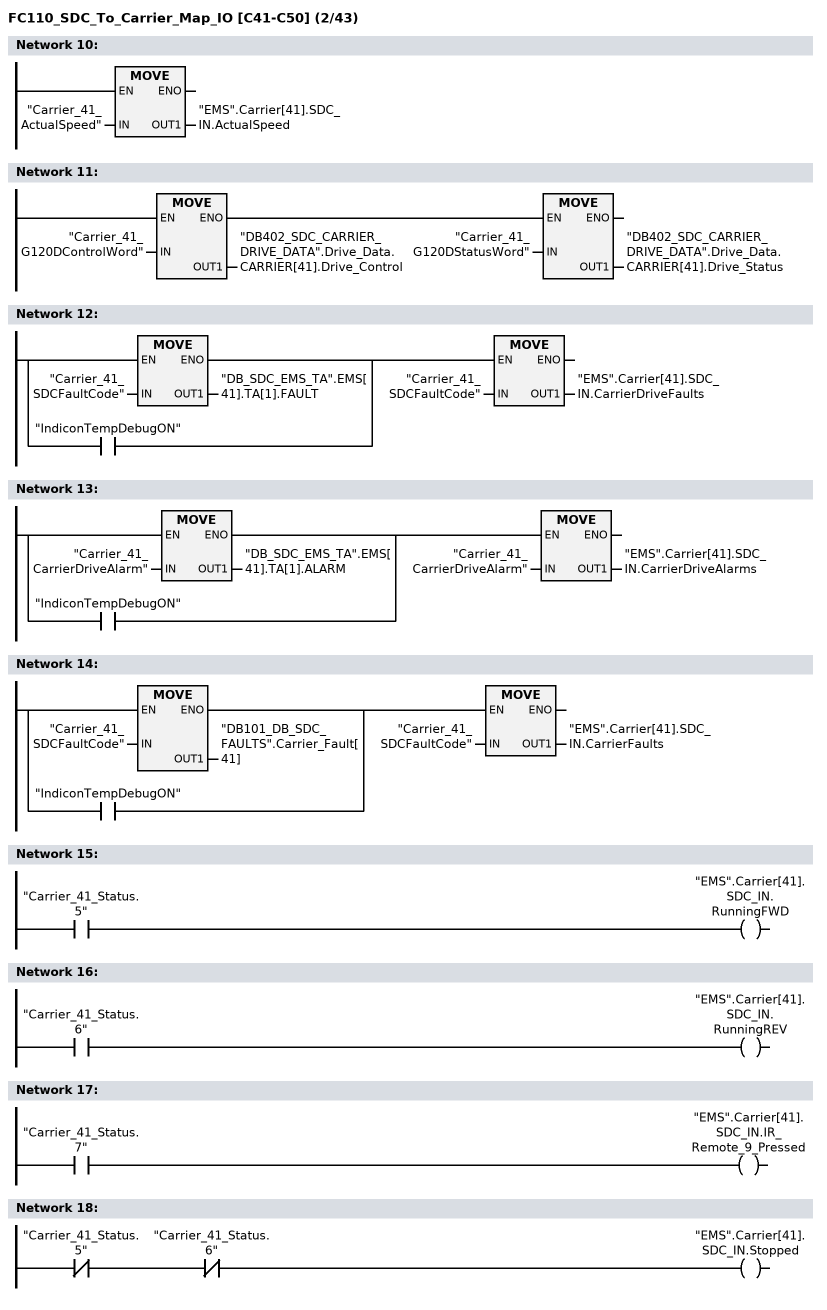
   RUNG wire#powerrail
      Move(in := "Carrier_41_ActualSpeed", out1 => "EMS".Carrier[41].SDC_IN.ActualSpeed)
   END_RUNG
   // the same network as SCL:
   "EMS".Carrier[41].SDC_IN.ActualSpeed := "Carrier_41_ActualSpeed";
END_REGION

REGION Network 11
   RUNG wire#powerrail
      Move(in := "Carrier_41_G120DControlWord", out1 => "DB402_SDC_CARRIER_DRIVE_DATA".Drive_Data.CARRIER[41].Drive_Control)
      Move(in := "Carrier_41_G120DStatusWord", out1 => "DB402_SDC_CARRIER_DRIVE_DATA".Drive_Data.CARRIER[41].Drive_Status)
   END_RUNG
   // the same network as SCL:
   "DB402_SDC_CARRIER_DRIVE_DATA".Drive_Data.CARRIER[41].Drive_Control := "Carrier_41_G120DControlWord";
   "DB402_SDC_CARRIER_DRIVE_DATA".Drive_Data.CARRIER[41].Drive_Status := "Carrier_41_G120DStatusWord";
END_REGION

REGION Network 12
   RUNG wire#powerrail
      Move(in := "Carrier_41_SDCFaultCode", out1 => "DB_SDC_EMS_TA".EMS[41].TA[1].FAULT)
      wire#w1
      Move(in := "Carrier_41_SDCFaultCode", out1 => "EMS".Carrier[41].SDC_IN.CarrierDriveFaults)
   END_RUNG
   RUNG wire#powerrail
      Contact( "IndiconTempDebugON" )
   END_RUNG wire#w1
   // the same network as SCL:
   "DB_SDC_EMS_TA".EMS[41].TA[1].FAULT := "Carrier_41_SDCFaultCode";
   IF TRUE OR "IndiconTempDebugON" THEN
       "EMS".Carrier[41].SDC_IN.CarrierDriveFaults := "Carrier_41_SDCFaultCode";
   END_IF;
END_REGION

REGION Network 13
   RUNG wire#powerrail
      Move(in := "Carrier_41_CarrierDriveAlarm", out1 => "DB_SDC_EMS_TA".EMS[41].TA[1].ALARM)
      wire#w1
      Move(in := "Carrier_41_CarrierDriveAlarm", out1 => "EMS".Carrier[41].SDC_IN.CarrierDriveAlarms)
   END_RUNG
   RUNG wire#powerrail
      Contact( "IndiconTempDebugON" )
   END_RUNG wire#w1
   // the same network as SCL:
   "DB_SDC_EMS_TA".EMS[41].TA[1].ALARM := "Carrier_41_CarrierDriveAlarm";
   IF TRUE OR "IndiconTempDebugON" THEN
       "EMS".Carrier[41].SDC_IN.CarrierDriveAlarms := "Carrier_41_CarrierDriveAlarm";
   END_IF;
END_REGION

REGION Network 14
   RUNG wire#powerrail
      Move(in := "Carrier_41_SDCFaultCode", out1 => "DB101_DB_SDC_FAULTS".Carrier_Fault[41])
      wire#w1
      Move(in := "Carrier_41_SDCFaultCode", out1 => "EMS".Carrier[41].SDC_IN.CarrierFaults)
   END_RUNG
   RUNG wire#powerrail
      Contact( "IndiconTempDebugON" )
   END_RUNG wire#w1
   // the same network as SCL:
   "DB101_DB_SDC_FAULTS".Carrier_Fault[41] := "Carrier_41_SDCFaultCode";
   IF TRUE OR "IndiconTempDebugON" THEN
       "EMS".Carrier[41].SDC_IN.CarrierFaults := "Carrier_41_SDCFaultCode";
   END_IF;
END_REGION

REGION Network 15
   RUNG wire#powerrail
      Contact( "Carrier_41_Status.5" )
      Coil( "EMS".Carrier[41].SDC_IN.RunningFWD )
   END_RUNG
   // the same network as SCL:
   "EMS".Carrier[41].SDC_IN.RunningFWD := "Carrier_41_Status.5";
END_REGION

REGION Network 16
   RUNG wire#powerrail
      Contact( "Carrier_41_Status.6" )
      Coil( "EMS".Carrier[41].SDC_IN.RunningREV )
   END_RUNG
   // the same network as SCL:
   "EMS".Carrier[41].SDC_IN.RunningREV := "Carrier_41_Status.6";
END_REGION

REGION Network 17
   RUNG wire#powerrail
      Contact( "Carrier_41_Status.7" )
      Coil( "EMS".Carrier[41].SDC_IN.IR_Remote_9_Pressed )
   END_RUNG
   // the same network as SCL:
   "EMS".Carrier[41].SDC_IN.IR_Remote_9_Pressed := "Carrier_41_Status.7";
END_REGION

REGION Network 18
   RUNG wire#powerrail
      I_Contact( "Carrier_41_Status.5" )
      I_Contact( "Carrier_41_Status.6" )
      Coil( "EMS".Carrier[41].SDC_IN.Stopped )
   END_RUNG
   // the same network as SCL:
   "EMS".Carrier[41].SDC_IN.Stopped := NOT "Carrier_41_Status.5" AND NOT "Carrier_41_Status.6";
END_REGION

REGION Network 19
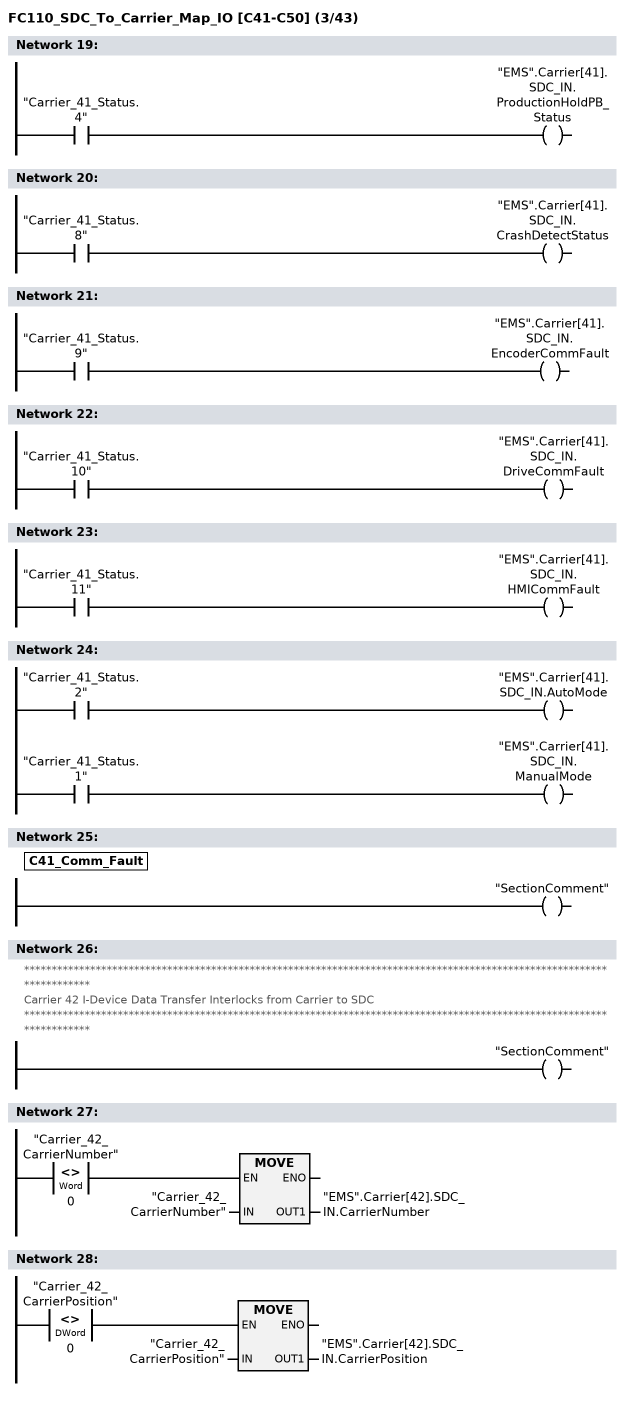
   RUNG wire#powerrail
      Contact( "Carrier_41_Status.4" )
      Coil( "EMS".Carrier[41].SDC_IN.ProductionHoldPB_Status )
   END_RUNG
   // the same network as SCL:
   "EMS".Carrier[41].SDC_IN.ProductionHoldPB_Status := "Carrier_41_Status.4";
END_REGION

REGION Network 20
   RUNG wire#powerrail
      Contact( "Carrier_41_Status.8" )
      Coil( "EMS".Carrier[41].SDC_IN.CrashDetectStatus )
   END_RUNG
   // the same network as SCL:
   "EMS".Carrier[41].SDC_IN.CrashDetectStatus := "Carrier_41_Status.8";
END_REGION

REGION Network 21
   RUNG wire#powerrail
      Contact( "Carrier_41_Status.9" )
      Coil( "EMS".Carrier[41].SDC_IN.EncoderCommFault )
   END_RUNG
   // the same network as SCL:
   "EMS".Carrier[41].SDC_IN.EncoderCommFault := "Carrier_41_Status.9";
END_REGION

REGION Network 22
   RUNG wire#powerrail
      Contact( "Carrier_41_Status.10" )
      Coil( "EMS".Carrier[41].SDC_IN.DriveCommFault )
   END_RUNG
   // the same network as SCL:
   "EMS".Carrier[41].SDC_IN.DriveCommFault := "Carrier_41_Status.10";
END_REGION

REGION Network 23
   RUNG wire#powerrail
      Contact( "Carrier_41_Status.11" )
      Coil( "EMS".Carrier[41].SDC_IN.HMICommFault )
   END_RUNG
   // the same network as SCL:
   "EMS".Carrier[41].SDC_IN.HMICommFault := "Carrier_41_Status.11";
END_REGION

REGION Network 24
   RUNG wire#powerrail
      Contact( "Carrier_41_Status.2" )
      Coil( "EMS".Carrier[41].SDC_IN.AutoMode )
   END_RUNG
   RUNG wire#powerrail
      Contact( "Carrier_41_Status.1" )
      Coil( "EMS".Carrier[41].SDC_IN.ManualMode )
   END_RUNG
   // the same network as SCL:
   "EMS".Carrier[41].SDC_IN.AutoMode := "Carrier_41_Status.2";
   "EMS".Carrier[41].SDC_IN.ManualMode := "Carrier_41_Status.1";
END_REGION

REGION Network 25
   Label( C41_Comm_Fault )
   RUNG wire#powerrail
      Coil( "SectionComment" )
   END_RUNG
   // the same network as SCL:
   C41_Comm_Fault:
   "SectionComment" := TRUE;
END_REGION

REGION Network 26
   // **********************************************************************************************************************
   // 
   // Carrier 42 I-Device Data Transfer Interlocks from Carrier to SDC
   // 
   // **********************************************************************************************************************
   RUNG wire#powerrail
      Coil( "SectionComment" )
   END_RUNG
   // the same network as SCL:
   "SectionComment" := TRUE;
END_REGION

REGION Network 27
   RUNG wire#powerrail
      { S7_Templates := "SrcType := Word" } NE_Contact(in1 := "Carrier_42_CarrierNumber", in2 := 0)
      Move(in := "Carrier_42_CarrierNumber", out1 => "EMS".Carrier[42].SDC_IN.CarrierNumber)
   END_RUNG
   // the same network as SCL:
   IF "Carrier_42_CarrierNumber" <> 0 THEN
       "EMS".Carrier[42].SDC_IN.CarrierNumber := "Carrier_42_CarrierNumber";
   END_IF;
END_REGION

REGION Network 28
   RUNG wire#powerrail
      { S7_Templates := "SrcType := DWord" } NE_Contact(in1 := "Carrier_42_CarrierPosition", in2 := 0)
      Move(in := "Carrier_42_CarrierPosition", out1 => "EMS".Carrier[42].SDC_IN.CarrierPosition)
   END_RUNG
   // the same network as SCL:
   IF "Carrier_42_CarrierPosition" <> 0 THEN
       "EMS".Carrier[42].SDC_IN.CarrierPosition := "Carrier_42_CarrierPosition";
   END_IF;
END_REGION

REGION Network 29
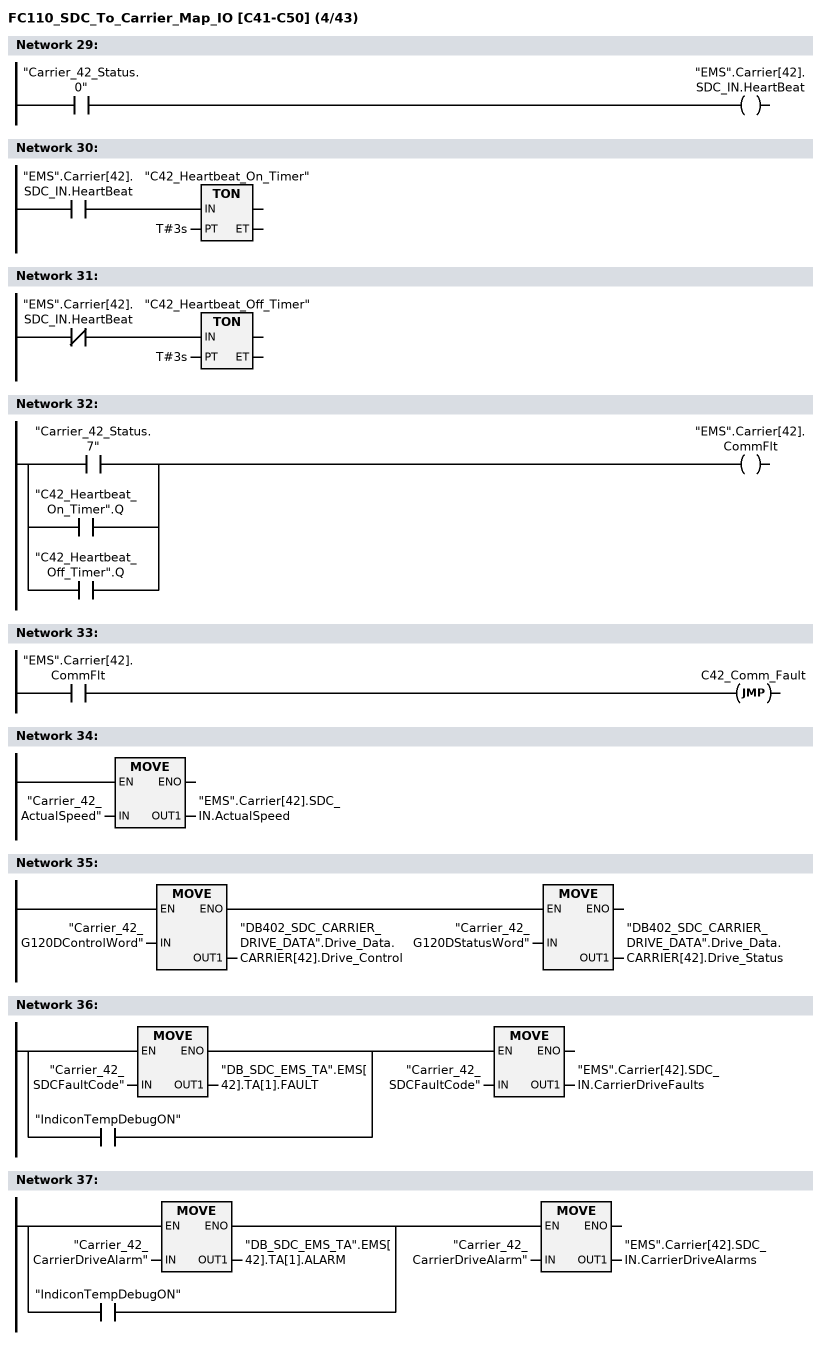
   RUNG wire#powerrail
      Contact( "Carrier_42_Status.0" )
      Coil( "EMS".Carrier[42].SDC_IN.HeartBeat )
   END_RUNG
   // the same network as SCL:
   "EMS".Carrier[42].SDC_IN.HeartBeat := "Carrier_42_Status.0";
END_REGION

REGION Network 30
   "C42_Heartbeat_On_Timer".TON(IN := "EMS".Carrier[42].SDC_IN.HeartBeat, PT := T#3s);
END_REGION

REGION Network 31
   "C42_Heartbeat_Off_Timer".TON(IN := NOT "EMS".Carrier[42].SDC_IN.HeartBeat, PT := T#3s);
END_REGION

REGION Network 32
   RUNG wire#powerrail
      Contact( "Carrier_42_Status.7" )
      wire#w1
      Coil( "EMS".Carrier[42].CommFlt )
   END_RUNG
   RUNG wire#powerrail
      Contact( "C42_Heartbeat_On_Timer".Q )
   END_RUNG wire#w1
   RUNG wire#powerrail
      Contact( "C42_Heartbeat_Off_Timer".Q )
   END_RUNG wire#w1
   // the same network as SCL:
   "EMS".Carrier[42].CommFlt := "Carrier_42_Status.7" OR "C42_Heartbeat_On_Timer".Q OR "C42_Heartbeat_Off_Timer".Q;
END_REGION

REGION Network 33
   RUNG wire#powerrail
      Contact( "EMS".Carrier[42].CommFlt )
      JumpCoil( C42_Comm_Fault )
   END_RUNG
   // the same network as SCL:
   IF "EMS".Carrier[42].CommFlt THEN GOTO C42_Comm_Fault; END_IF;
END_REGION

REGION Network 34
   RUNG wire#powerrail
      Move(in := "Carrier_42_ActualSpeed", out1 => "EMS".Carrier[42].SDC_IN.ActualSpeed)
   END_RUNG
   // the same network as SCL:
   "EMS".Carrier[42].SDC_IN.ActualSpeed := "Carrier_42_ActualSpeed";
END_REGION

REGION Network 35
   RUNG wire#powerrail
      Move(in := "Carrier_42_G120DControlWord", out1 => "DB402_SDC_CARRIER_DRIVE_DATA".Drive_Data.CARRIER[42].Drive_Control)
      Move(in := "Carrier_42_G120DStatusWord", out1 => "DB402_SDC_CARRIER_DRIVE_DATA".Drive_Data.CARRIER[42].Drive_Status)
   END_RUNG
   // the same network as SCL:
   "DB402_SDC_CARRIER_DRIVE_DATA".Drive_Data.CARRIER[42].Drive_Control := "Carrier_42_G120DControlWord";
   "DB402_SDC_CARRIER_DRIVE_DATA".Drive_Data.CARRIER[42].Drive_Status := "Carrier_42_G120DStatusWord";
END_REGION

REGION Network 36
   RUNG wire#powerrail
      Move(in := "Carrier_42_SDCFaultCode", out1 => "DB_SDC_EMS_TA".EMS[42].TA[1].FAULT)
      wire#w1
      Move(in := "Carrier_42_SDCFaultCode", out1 => "EMS".Carrier[42].SDC_IN.CarrierDriveFaults)
   END_RUNG
   RUNG wire#powerrail
      Contact( "IndiconTempDebugON" )
   END_RUNG wire#w1
   // the same network as SCL:
   "DB_SDC_EMS_TA".EMS[42].TA[1].FAULT := "Carrier_42_SDCFaultCode";
   IF TRUE OR "IndiconTempDebugON" THEN
       "EMS".Carrier[42].SDC_IN.CarrierDriveFaults := "Carrier_42_SDCFaultCode";
   END_IF;
END_REGION

REGION Network 37
   RUNG wire#powerrail
      Move(in := "Carrier_42_CarrierDriveAlarm", out1 => "DB_SDC_EMS_TA".EMS[42].TA[1].ALARM)
      wire#w1
      Move(in := "Carrier_42_CarrierDriveAlarm", out1 => "EMS".Carrier[42].SDC_IN.CarrierDriveAlarms)
   END_RUNG
   RUNG wire#powerrail
      Contact( "IndiconTempDebugON" )
   END_RUNG wire#w1
   // the same network as SCL:
   "DB_SDC_EMS_TA".EMS[42].TA[1].ALARM := "Carrier_42_CarrierDriveAlarm";
   IF TRUE OR "IndiconTempDebugON" THEN
       "EMS".Carrier[42].SDC_IN.CarrierDriveAlarms := "Carrier_42_CarrierDriveAlarm";
   END_IF;
END_REGION

REGION Network 38
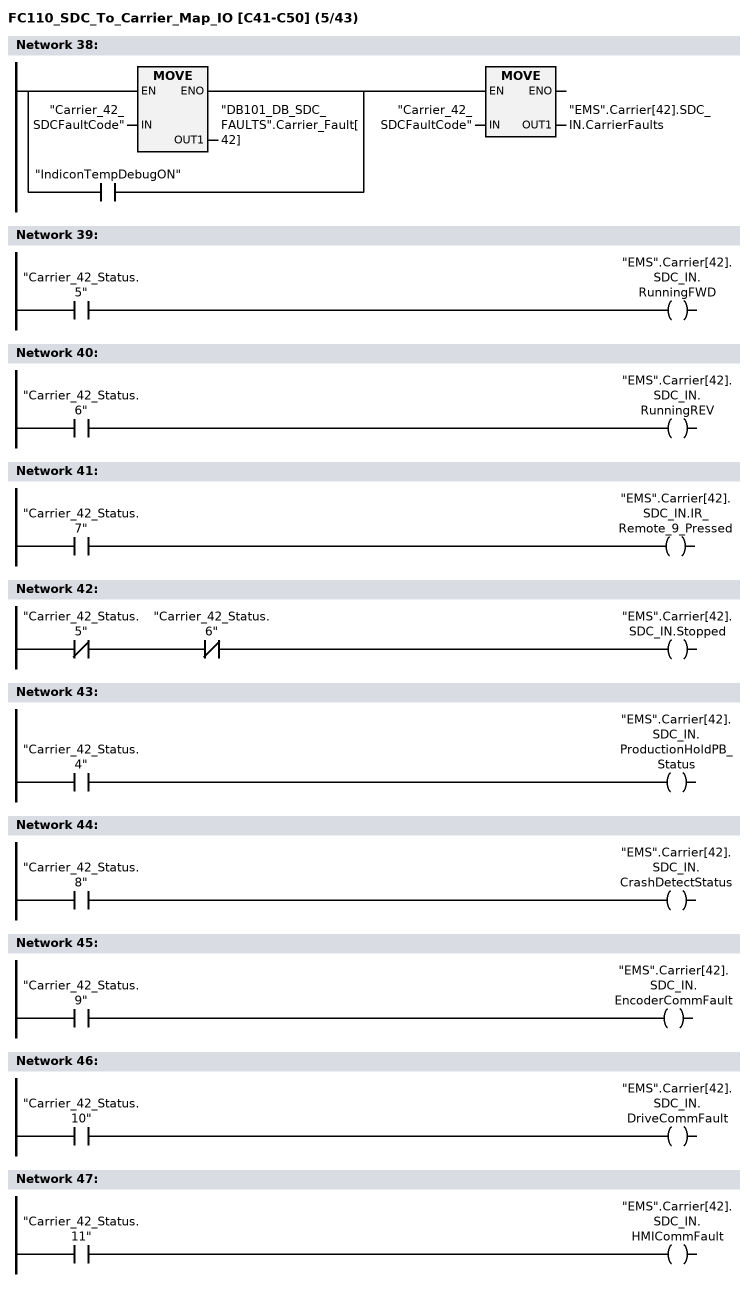
   RUNG wire#powerrail
      Move(in := "Carrier_42_SDCFaultCode", out1 => "DB101_DB_SDC_FAULTS".Carrier_Fault[42])
      wire#w1
      Move(in := "Carrier_42_SDCFaultCode", out1 => "EMS".Carrier[42].SDC_IN.CarrierFaults)
   END_RUNG
   RUNG wire#powerrail
      Contact( "IndiconTempDebugON" )
   END_RUNG wire#w1
   // the same network as SCL:
   "DB101_DB_SDC_FAULTS".Carrier_Fault[42] := "Carrier_42_SDCFaultCode";
   IF TRUE OR "IndiconTempDebugON" THEN
       "EMS".Carrier[42].SDC_IN.CarrierFaults := "Carrier_42_SDCFaultCode";
   END_IF;
END_REGION

REGION Network 39
   RUNG wire#powerrail
      Contact( "Carrier_42_Status.5" )
      Coil( "EMS".Carrier[42].SDC_IN.RunningFWD )
   END_RUNG
   // the same network as SCL:
   "EMS".Carrier[42].SDC_IN.RunningFWD := "Carrier_42_Status.5";
END_REGION

REGION Network 40
   RUNG wire#powerrail
      Contact( "Carrier_42_Status.6" )
      Coil( "EMS".Carrier[42].SDC_IN.RunningREV )
   END_RUNG
   // the same network as SCL:
   "EMS".Carrier[42].SDC_IN.RunningREV := "Carrier_42_Status.6";
END_REGION

REGION Network 41
   RUNG wire#powerrail
      Contact( "Carrier_42_Status.7" )
      Coil( "EMS".Carrier[42].SDC_IN.IR_Remote_9_Pressed )
   END_RUNG
   // the same network as SCL:
   "EMS".Carrier[42].SDC_IN.IR_Remote_9_Pressed := "Carrier_42_Status.7";
END_REGION

REGION Network 42
   RUNG wire#powerrail
      I_Contact( "Carrier_42_Status.5" )
      I_Contact( "Carrier_42_Status.6" )
      Coil( "EMS".Carrier[42].SDC_IN.Stopped )
   END_RUNG
   // the same network as SCL:
   "EMS".Carrier[42].SDC_IN.Stopped := NOT "Carrier_42_Status.5" AND NOT "Carrier_42_Status.6";
END_REGION

REGION Network 43
   RUNG wire#powerrail
      Contact( "Carrier_42_Status.4" )
      Coil( "EMS".Carrier[42].SDC_IN.ProductionHoldPB_Status )
   END_RUNG
   // the same network as SCL:
   "EMS".Carrier[42].SDC_IN.ProductionHoldPB_Status := "Carrier_42_Status.4";
END_REGION

REGION Network 44
   RUNG wire#powerrail
      Contact( "Carrier_42_Status.8" )
      Coil( "EMS".Carrier[42].SDC_IN.CrashDetectStatus )
   END_RUNG
   // the same network as SCL:
   "EMS".Carrier[42].SDC_IN.CrashDetectStatus := "Carrier_42_Status.8";
END_REGION

REGION Network 45
   RUNG wire#powerrail
      Contact( "Carrier_42_Status.9" )
      Coil( "EMS".Carrier[42].SDC_IN.EncoderCommFault )
   END_RUNG
   // the same network as SCL:
   "EMS".Carrier[42].SDC_IN.EncoderCommFault := "Carrier_42_Status.9";
END_REGION

REGION Network 46
   RUNG wire#powerrail
      Contact( "Carrier_42_Status.10" )
      Coil( "EMS".Carrier[42].SDC_IN.DriveCommFault )
   END_RUNG
   // the same network as SCL:
   "EMS".Carrier[42].SDC_IN.DriveCommFault := "Carrier_42_Status.10";
END_REGION

REGION Network 47
   RUNG wire#powerrail
      Contact( "Carrier_42_Status.11" )
      Coil( "EMS".Carrier[42].SDC_IN.HMICommFault )
   END_RUNG
   // the same network as SCL:
   "EMS".Carrier[42].SDC_IN.HMICommFault := "Carrier_42_Status.11";
END_REGION

REGION Network 48
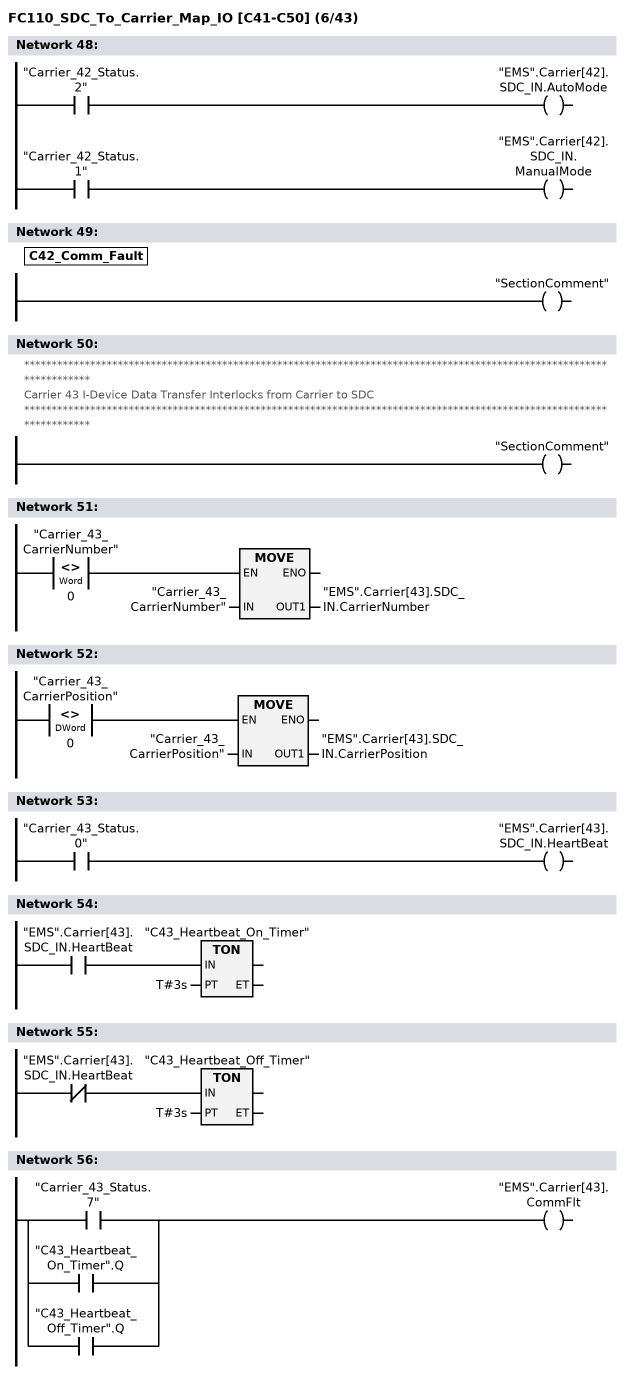
   RUNG wire#powerrail
      Contact( "Carrier_42_Status.2" )
      Coil( "EMS".Carrier[42].SDC_IN.AutoMode )
   END_RUNG
   RUNG wire#powerrail
      Contact( "Carrier_42_Status.1" )
      Coil( "EMS".Carrier[42].SDC_IN.ManualMode )
   END_RUNG
   // the same network as SCL:
   "EMS".Carrier[42].SDC_IN.AutoMode := "Carrier_42_Status.2";
   "EMS".Carrier[42].SDC_IN.ManualMode := "Carrier_42_Status.1";
END_REGION

REGION Network 49
   Label( C42_Comm_Fault )
   RUNG wire#powerrail
      Coil( "SectionComment" )
   END_RUNG
   // the same network as SCL:
   C42_Comm_Fault:
   "SectionComment" := TRUE;
END_REGION

REGION Network 50
   // **********************************************************************************************************************
   // 
   // Carrier 43 I-Device Data Transfer Interlocks from Carrier to SDC
   // 
   // **********************************************************************************************************************
   RUNG wire#powerrail
      Coil( "SectionComment" )
   END_RUNG
   // the same network as SCL:
   "SectionComment" := TRUE;
END_REGION

REGION Network 51
   RUNG wire#powerrail
      { S7_Templates := "SrcType := Word" } NE_Contact(in1 := "Carrier_43_CarrierNumber", in2 := 0)
      Move(in := "Carrier_43_CarrierNumber", out1 => "EMS".Carrier[43].SDC_IN.CarrierNumber)
   END_RUNG
   // the same network as SCL:
   IF "Carrier_43_CarrierNumber" <> 0 THEN
       "EMS".Carrier[43].SDC_IN.CarrierNumber := "Carrier_43_CarrierNumber";
   END_IF;
END_REGION

REGION Network 52
   RUNG wire#powerrail
      { S7_Templates := "SrcType := DWord" } NE_Contact(in1 := "Carrier_43_CarrierPosition", in2 := 0)
      Move(in := "Carrier_43_CarrierPosition", out1 => "EMS".Carrier[43].SDC_IN.CarrierPosition)
   END_RUNG
   // the same network as SCL:
   IF "Carrier_43_CarrierPosition" <> 0 THEN
       "EMS".Carrier[43].SDC_IN.CarrierPosition := "Carrier_43_CarrierPosition";
   END_IF;
END_REGION

REGION Network 53
   RUNG wire#powerrail
      Contact( "Carrier_43_Status.0" )
      Coil( "EMS".Carrier[43].SDC_IN.HeartBeat )
   END_RUNG
   // the same network as SCL:
   "EMS".Carrier[43].SDC_IN.HeartBeat := "Carrier_43_Status.0";
END_REGION

REGION Network 54
   "C43_Heartbeat_On_Timer".TON(IN := "EMS".Carrier[43].SDC_IN.HeartBeat, PT := T#3s);
END_REGION

REGION Network 55
   "C43_Heartbeat_Off_Timer".TON(IN := NOT "EMS".Carrier[43].SDC_IN.HeartBeat, PT := T#3s);
END_REGION

REGION Network 56
   RUNG wire#powerrail
      Contact( "Carrier_43_Status.7" )
      wire#w1
      Coil( "EMS".Carrier[43].CommFlt )
   END_RUNG
   RUNG wire#powerrail
      Contact( "C43_Heartbeat_On_Timer".Q )
   END_RUNG wire#w1
   RUNG wire#powerrail
      Contact( "C43_Heartbeat_Off_Timer".Q )
   END_RUNG wire#w1
   // the same network as SCL:
   "EMS".Carrier[43].CommFlt := "Carrier_43_Status.7" OR "C43_Heartbeat_On_Timer".Q OR "C43_Heartbeat_Off_Timer".Q;
END_REGION

REGION Network 57
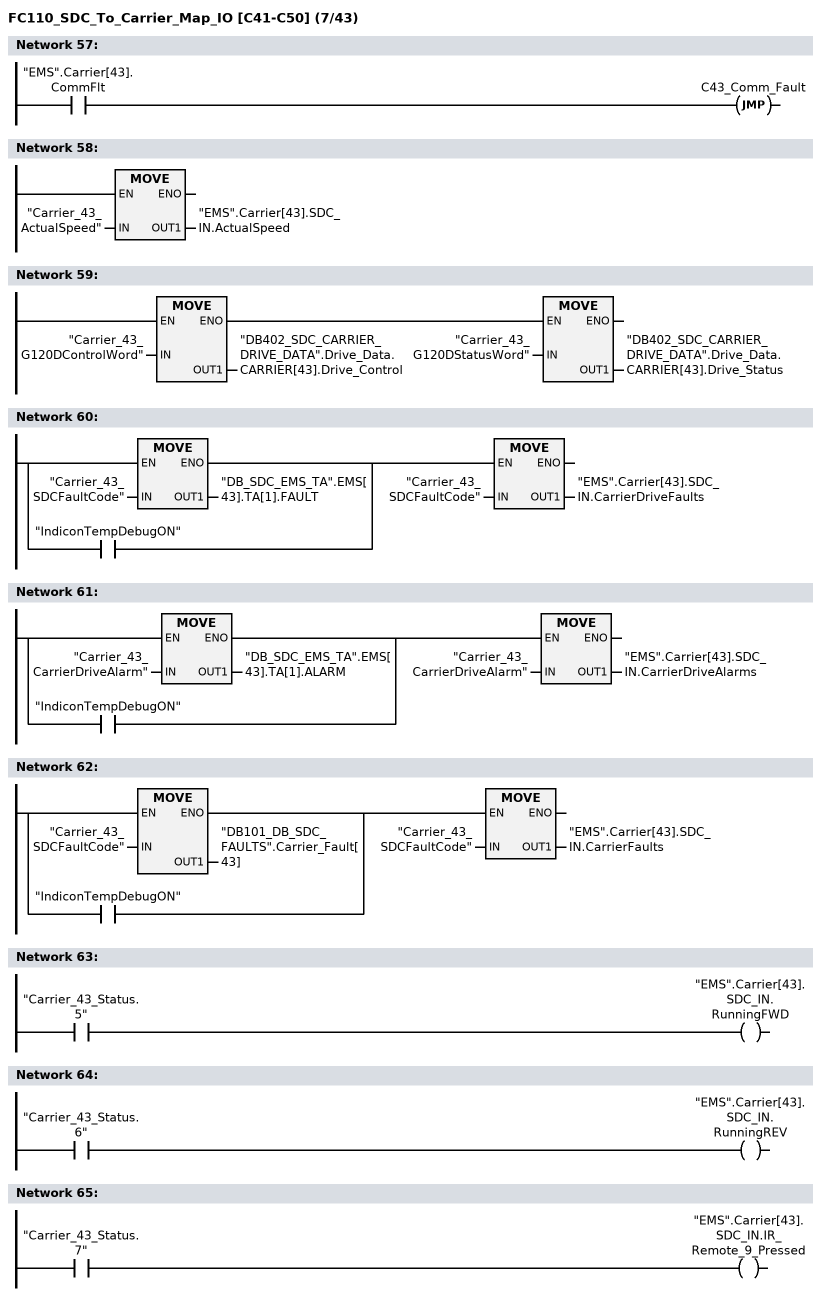
   RUNG wire#powerrail
      Contact( "EMS".Carrier[43].CommFlt )
      JumpCoil( C43_Comm_Fault )
   END_RUNG
   // the same network as SCL:
   IF "EMS".Carrier[43].CommFlt THEN GOTO C43_Comm_Fault; END_IF;
END_REGION

REGION Network 58
   RUNG wire#powerrail
      Move(in := "Carrier_43_ActualSpeed", out1 => "EMS".Carrier[43].SDC_IN.ActualSpeed)
   END_RUNG
   // the same network as SCL:
   "EMS".Carrier[43].SDC_IN.ActualSpeed := "Carrier_43_ActualSpeed";
END_REGION

REGION Network 59
   RUNG wire#powerrail
      Move(in := "Carrier_43_G120DControlWord", out1 => "DB402_SDC_CARRIER_DRIVE_DATA".Drive_Data.CARRIER[43].Drive_Control)
      Move(in := "Carrier_43_G120DStatusWord", out1 => "DB402_SDC_CARRIER_DRIVE_DATA".Drive_Data.CARRIER[43].Drive_Status)
   END_RUNG
   // the same network as SCL:
   "DB402_SDC_CARRIER_DRIVE_DATA".Drive_Data.CARRIER[43].Drive_Control := "Carrier_43_G120DControlWord";
   "DB402_SDC_CARRIER_DRIVE_DATA".Drive_Data.CARRIER[43].Drive_Status := "Carrier_43_G120DStatusWord";
END_REGION

REGION Network 60
   RUNG wire#powerrail
      Move(in := "Carrier_43_SDCFaultCode", out1 => "DB_SDC_EMS_TA".EMS[43].TA[1].FAULT)
      wire#w1
      Move(in := "Carrier_43_SDCFaultCode", out1 => "EMS".Carrier[43].SDC_IN.CarrierDriveFaults)
   END_RUNG
   RUNG wire#powerrail
      Contact( "IndiconTempDebugON" )
   END_RUNG wire#w1
   // the same network as SCL:
   "DB_SDC_EMS_TA".EMS[43].TA[1].FAULT := "Carrier_43_SDCFaultCode";
   IF TRUE OR "IndiconTempDebugON" THEN
       "EMS".Carrier[43].SDC_IN.CarrierDriveFaults := "Carrier_43_SDCFaultCode";
   END_IF;
END_REGION

REGION Network 61
   RUNG wire#powerrail
      Move(in := "Carrier_43_CarrierDriveAlarm", out1 => "DB_SDC_EMS_TA".EMS[43].TA[1].ALARM)
      wire#w1
      Move(in := "Carrier_43_CarrierDriveAlarm", out1 => "EMS".Carrier[43].SDC_IN.CarrierDriveAlarms)
   END_RUNG
   RUNG wire#powerrail
      Contact( "IndiconTempDebugON" )
   END_RUNG wire#w1
   // the same network as SCL:
   "DB_SDC_EMS_TA".EMS[43].TA[1].ALARM := "Carrier_43_CarrierDriveAlarm";
   IF TRUE OR "IndiconTempDebugON" THEN
       "EMS".Carrier[43].SDC_IN.CarrierDriveAlarms := "Carrier_43_CarrierDriveAlarm";
   END_IF;
END_REGION

REGION Network 62
   RUNG wire#powerrail
      Move(in := "Carrier_43_SDCFaultCode", out1 => "DB101_DB_SDC_FAULTS".Carrier_Fault[43])
      wire#w1
      Move(in := "Carrier_43_SDCFaultCode", out1 => "EMS".Carrier[43].SDC_IN.CarrierFaults)
   END_RUNG
   RUNG wire#powerrail
      Contact( "IndiconTempDebugON" )
   END_RUNG wire#w1
   // the same network as SCL:
   "DB101_DB_SDC_FAULTS".Carrier_Fault[43] := "Carrier_43_SDCFaultCode";
   IF TRUE OR "IndiconTempDebugON" THEN
       "EMS".Carrier[43].SDC_IN.CarrierFaults := "Carrier_43_SDCFaultCode";
   END_IF;
END_REGION

REGION Network 63
   RUNG wire#powerrail
      Contact( "Carrier_43_Status.5" )
      Coil( "EMS".Carrier[43].SDC_IN.RunningFWD )
   END_RUNG
   // the same network as SCL:
   "EMS".Carrier[43].SDC_IN.RunningFWD := "Carrier_43_Status.5";
END_REGION

REGION Network 64
   RUNG wire#powerrail
      Contact( "Carrier_43_Status.6" )
      Coil( "EMS".Carrier[43].SDC_IN.RunningREV )
   END_RUNG
   // the same network as SCL:
   "EMS".Carrier[43].SDC_IN.RunningREV := "Carrier_43_Status.6";
END_REGION

REGION Network 65
   RUNG wire#powerrail
      Contact( "Carrier_43_Status.7" )
      Coil( "EMS".Carrier[43].SDC_IN.IR_Remote_9_Pressed )
   END_RUNG
   // the same network as SCL:
   "EMS".Carrier[43].SDC_IN.IR_Remote_9_Pressed := "Carrier_43_Status.7";
END_REGION

REGION Network 66
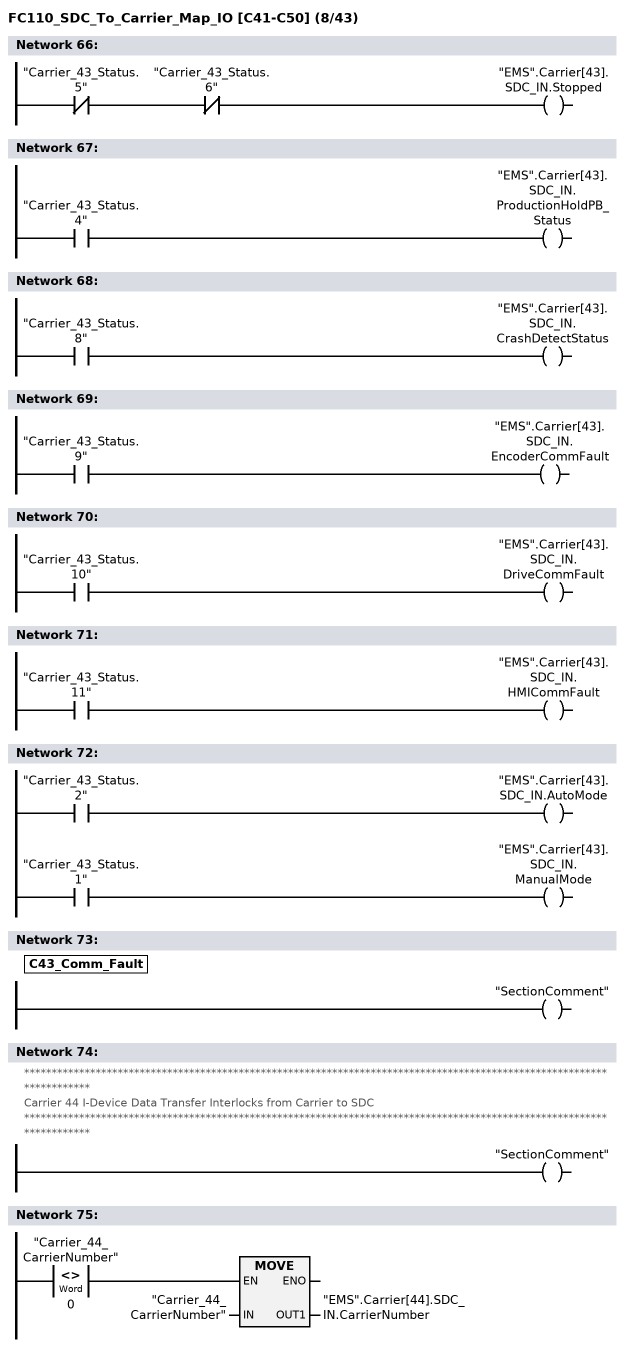
   RUNG wire#powerrail
      I_Contact( "Carrier_43_Status.5" )
      I_Contact( "Carrier_43_Status.6" )
      Coil( "EMS".Carrier[43].SDC_IN.Stopped )
   END_RUNG
   // the same network as SCL:
   "EMS".Carrier[43].SDC_IN.Stopped := NOT "Carrier_43_Status.5" AND NOT "Carrier_43_Status.6";
END_REGION

REGION Network 67
   RUNG wire#powerrail
      Contact( "Carrier_43_Status.4" )
      Coil( "EMS".Carrier[43].SDC_IN.ProductionHoldPB_Status )
   END_RUNG
   // the same network as SCL:
   "EMS".Carrier[43].SDC_IN.ProductionHoldPB_Status := "Carrier_43_Status.4";
END_REGION

REGION Network 68
   RUNG wire#powerrail
      Contact( "Carrier_43_Status.8" )
      Coil( "EMS".Carrier[43].SDC_IN.CrashDetectStatus )
   END_RUNG
   // the same network as SCL:
   "EMS".Carrier[43].SDC_IN.CrashDetectStatus := "Carrier_43_Status.8";
END_REGION

REGION Network 69
   RUNG wire#powerrail
      Contact( "Carrier_43_Status.9" )
      Coil( "EMS".Carrier[43].SDC_IN.EncoderCommFault )
   END_RUNG
   // the same network as SCL:
   "EMS".Carrier[43].SDC_IN.EncoderCommFault := "Carrier_43_Status.9";
END_REGION

REGION Network 70
   RUNG wire#powerrail
      Contact( "Carrier_43_Status.10" )
      Coil( "EMS".Carrier[43].SDC_IN.DriveCommFault )
   END_RUNG
   // the same network as SCL:
   "EMS".Carrier[43].SDC_IN.DriveCommFault := "Carrier_43_Status.10";
END_REGION

REGION Network 71
   RUNG wire#powerrail
      Contact( "Carrier_43_Status.11" )
      Coil( "EMS".Carrier[43].SDC_IN.HMICommFault )
   END_RUNG
   // the same network as SCL:
   "EMS".Carrier[43].SDC_IN.HMICommFault := "Carrier_43_Status.11";
END_REGION

REGION Network 72
   RUNG wire#powerrail
      Contact( "Carrier_43_Status.2" )
      Coil( "EMS".Carrier[43].SDC_IN.AutoMode )
   END_RUNG
   RUNG wire#powerrail
      Contact( "Carrier_43_Status.1" )
      Coil( "EMS".Carrier[43].SDC_IN.ManualMode )
   END_RUNG
   // the same network as SCL:
   "EMS".Carrier[43].SDC_IN.AutoMode := "Carrier_43_Status.2";
   "EMS".Carrier[43].SDC_IN.ManualMode := "Carrier_43_Status.1";
END_REGION

REGION Network 73
   Label( C43_Comm_Fault )
   RUNG wire#powerrail
      Coil( "SectionComment" )
   END_RUNG
   // the same network as SCL:
   C43_Comm_Fault:
   "SectionComment" := TRUE;
END_REGION

REGION Network 74
   // **********************************************************************************************************************
   // 
   // Carrier 44 I-Device Data Transfer Interlocks from Carrier to SDC
   // 
   // **********************************************************************************************************************
   RUNG wire#powerrail
      Coil( "SectionComment" )
   END_RUNG
   // the same network as SCL:
   "SectionComment" := TRUE;
END_REGION

REGION Network 75
   RUNG wire#powerrail
      { S7_Templates := "SrcType := Word" } NE_Contact(in1 := "Carrier_44_CarrierNumber", in2 := 0)
      Move(in := "Carrier_44_CarrierNumber", out1 => "EMS".Carrier[44].SDC_IN.CarrierNumber)
   END_RUNG
   // the same network as SCL:
   IF "Carrier_44_CarrierNumber" <> 0 THEN
       "EMS".Carrier[44].SDC_IN.CarrierNumber := "Carrier_44_CarrierNumber";
   END_IF;
END_REGION

REGION Network 76
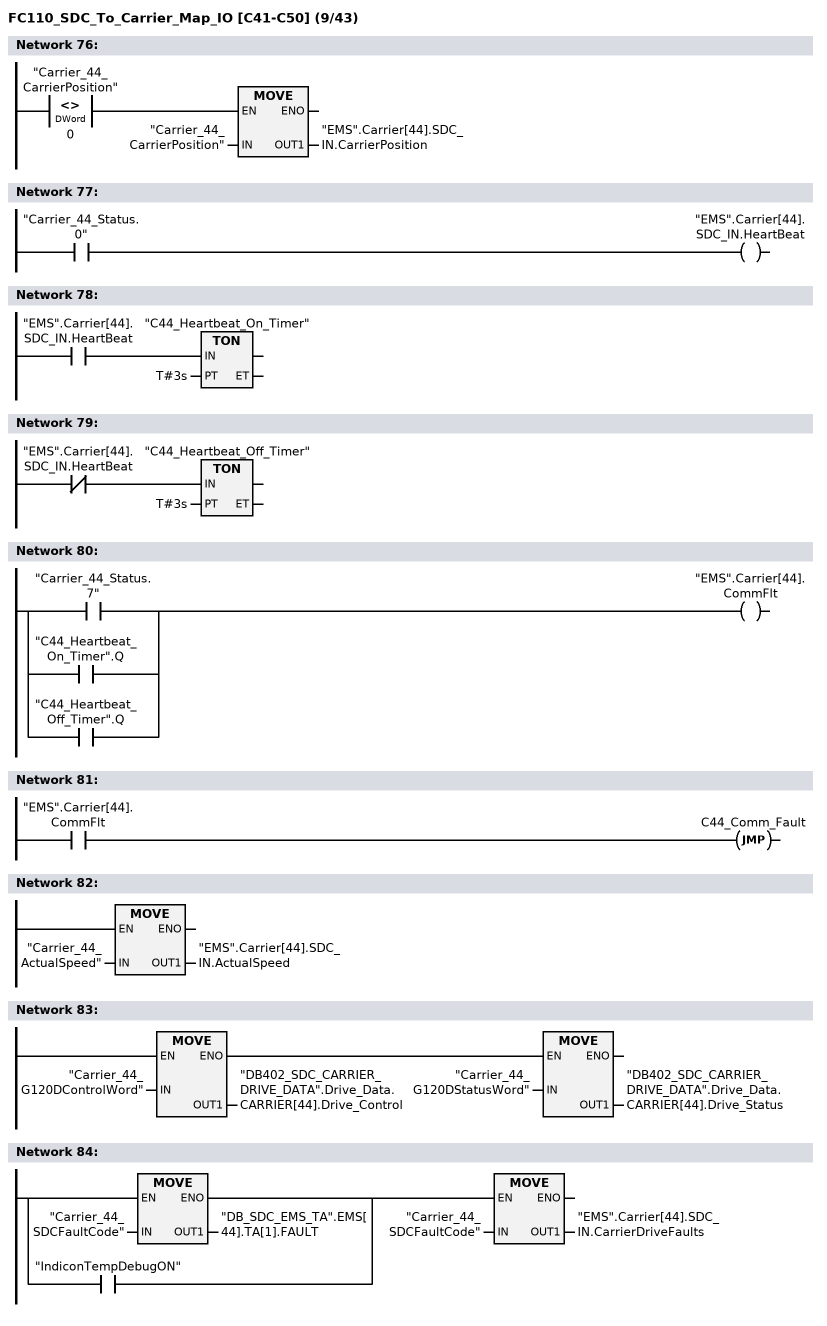
   RUNG wire#powerrail
      { S7_Templates := "SrcType := DWord" } NE_Contact(in1 := "Carrier_44_CarrierPosition", in2 := 0)
      Move(in := "Carrier_44_CarrierPosition", out1 => "EMS".Carrier[44].SDC_IN.CarrierPosition)
   END_RUNG
   // the same network as SCL:
   IF "Carrier_44_CarrierPosition" <> 0 THEN
       "EMS".Carrier[44].SDC_IN.CarrierPosition := "Carrier_44_CarrierPosition";
   END_IF;
END_REGION

REGION Network 77
   RUNG wire#powerrail
      Contact( "Carrier_44_Status.0" )
      Coil( "EMS".Carrier[44].SDC_IN.HeartBeat )
   END_RUNG
   // the same network as SCL:
   "EMS".Carrier[44].SDC_IN.HeartBeat := "Carrier_44_Status.0";
END_REGION

REGION Network 78
   "C44_Heartbeat_On_Timer".TON(IN := "EMS".Carrier[44].SDC_IN.HeartBeat, PT := T#3s);
END_REGION

REGION Network 79
   "C44_Heartbeat_Off_Timer".TON(IN := NOT "EMS".Carrier[44].SDC_IN.HeartBeat, PT := T#3s);
END_REGION

REGION Network 80
   RUNG wire#powerrail
      Contact( "Carrier_44_Status.7" )
      wire#w1
      Coil( "EMS".Carrier[44].CommFlt )
   END_RUNG
   RUNG wire#powerrail
      Contact( "C44_Heartbeat_On_Timer".Q )
   END_RUNG wire#w1
   RUNG wire#powerrail
      Contact( "C44_Heartbeat_Off_Timer".Q )
   END_RUNG wire#w1
   // the same network as SCL:
   "EMS".Carrier[44].CommFlt := "Carrier_44_Status.7" OR "C44_Heartbeat_On_Timer".Q OR "C44_Heartbeat_Off_Timer".Q;
END_REGION

REGION Network 81
   RUNG wire#powerrail
      Contact( "EMS".Carrier[44].CommFlt )
      JumpCoil( C44_Comm_Fault )
   END_RUNG
   // the same network as SCL:
   IF "EMS".Carrier[44].CommFlt THEN GOTO C44_Comm_Fault; END_IF;
END_REGION

REGION Network 82
   RUNG wire#powerrail
      Move(in := "Carrier_44_ActualSpeed", out1 => "EMS".Carrier[44].SDC_IN.ActualSpeed)
   END_RUNG
   // the same network as SCL:
   "EMS".Carrier[44].SDC_IN.ActualSpeed := "Carrier_44_ActualSpeed";
END_REGION
